REGION Network 164
   RUNG wire#powerrail
      Contact( "Carrier_27_Status.8" )
      Coil( "EMS".Carrier[27].SDC_IN.CrashDetectStatus )
   END_RUNG
   // the same network as SCL:
   "EMS".Carrier[27].SDC_IN.CrashDetectStatus := "Carrier_27_Status.8";
END_REGION

REGION Network 165
   RUNG wire#powerrail
      Contact( "Carrier_27_Status.9" )
      Coil( "EMS".Carrier[27].SDC_IN.EncoderCommFault )
   END_RUNG
   // the same network as SCL:
   "EMS".Carrier[27].SDC_IN.EncoderCommFault := "Carrier_27_Status.9";
END_REGION

REGION Network 166
   RUNG wire#powerrail
      Contact( "Carrier_27_Status.10" )
      Coil( "EMS".Carrier[27].SDC_IN.DriveCommFault )
   END_RUNG
   // the same network as SCL:
   "EMS".Carrier[27].SDC_IN.DriveCommFault := "Carrier_27_Status.10";
END_REGION

REGION Network 167
   RUNG wire#powerrail
      Contact( "Carrier_27_Status.11" )
      Coil( "EMS".Carrier[27].SDC_IN.HMICommFault )
   END_RUNG
   // the same network as SCL:
   "EMS".Carrier[27].SDC_IN.HMICommFault := "Carrier_27_Status.11";
END_REGION

REGION Network 168
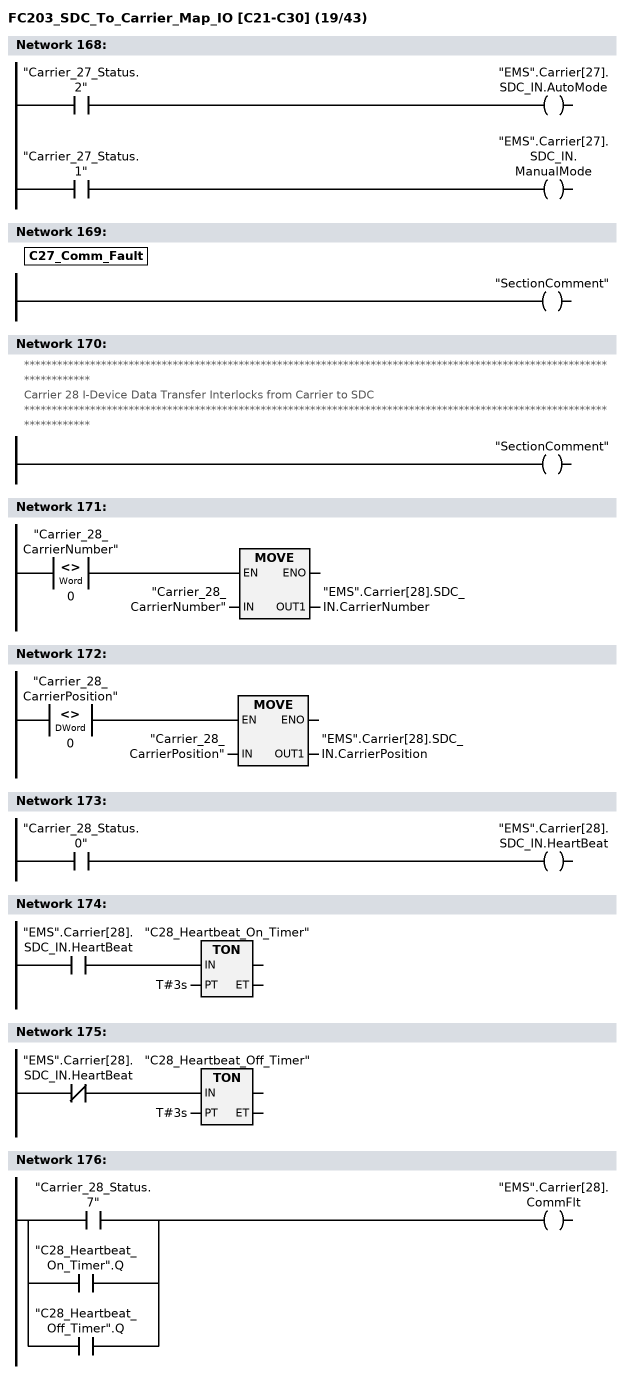
   RUNG wire#powerrail
      Contact( "Carrier_27_Status.2" )
      Coil( "EMS".Carrier[27].SDC_IN.AutoMode )
   END_RUNG
   RUNG wire#powerrail
      Contact( "Carrier_27_Status.1" )
      Coil( "EMS".Carrier[27].SDC_IN.ManualMode )
   END_RUNG
   // the same network as SCL:
   "EMS".Carrier[27].SDC_IN.AutoMode := "Carrier_27_Status.2";
   "EMS".Carrier[27].SDC_IN.ManualMode := "Carrier_27_Status.1";
END_REGION

REGION Network 169
   Label( C27_Comm_Fault )
   RUNG wire#powerrail
      Coil( "SectionComment" )
   END_RUNG
   // the same network as SCL:
   C27_Comm_Fault:
   "SectionComment" := TRUE;
END_REGION

REGION Network 170
   // **********************************************************************************************************************
   // 
   // Carrier 28 I-Device Data Transfer Interlocks from Carrier to SDC
   // 
   // **********************************************************************************************************************
   RUNG wire#powerrail
      Coil( "SectionComment" )
   END_RUNG
   // the same network as SCL:
   "SectionComment" := TRUE;
END_REGION

REGION Network 171
   RUNG wire#powerrail
      { S7_Templates := "SrcType := Word" } NE_Contact(in1 := "Carrier_28_CarrierNumber", in2 := 0)
      Move(in := "Carrier_28_CarrierNumber", out1 => "EMS".Carrier[28].SDC_IN.CarrierNumber)
   END_RUNG
   // the same network as SCL:
   IF "Carrier_28_CarrierNumber" <> 0 THEN
       "EMS".Carrier[28].SDC_IN.CarrierNumber := "Carrier_28_CarrierNumber";
   END_IF;
END_REGION

REGION Network 172
   RUNG wire#powerrail
      { S7_Templates := "SrcType := DWord" } NE_Contact(in1 := "Carrier_28_CarrierPosition", in2 := 0)
      Move(in := "Carrier_28_CarrierPosition", out1 => "EMS".Carrier[28].SDC_IN.CarrierPosition)
   END_RUNG
   // the same network as SCL:
   IF "Carrier_28_CarrierPosition" <> 0 THEN
       "EMS".Carrier[28].SDC_IN.CarrierPosition := "Carrier_28_CarrierPosition";
   END_IF;
END_REGION

REGION Network 173
   RUNG wire#powerrail
      Contact( "Carrier_28_Status.0" )
      Coil( "EMS".Carrier[28].SDC_IN.HeartBeat )
   END_RUNG
   // the same network as SCL:
   "EMS".Carrier[28].SDC_IN.HeartBeat := "Carrier_28_Status.0";
END_REGION

REGION Network 174
   "C28_Heartbeat_On_Timer".TON(IN := "EMS".Carrier[28].SDC_IN.HeartBeat, PT := T#3s);
END_REGION

REGION Network 175
   "C28_Heartbeat_Off_Timer".TON(IN := NOT "EMS".Carrier[28].SDC_IN.HeartBeat, PT := T#3s);
END_REGION

REGION Network 176
   RUNG wire#powerrail
      Contact( "Carrier_28_Status.7" )
      wire#w1
      Coil( "EMS".Carrier[28].CommFlt )
   END_RUNG
   RUNG wire#powerrail
      Contact( "C28_Heartbeat_On_Timer".Q )
   END_RUNG wire#w1
   RUNG wire#powerrail
      Contact( "C28_Heartbeat_Off_Timer".Q )
   END_RUNG wire#w1
   // the same network as SCL:
   "EMS".Carrier[28].CommFlt := "Carrier_28_Status.7" OR "C28_Heartbeat_On_Timer".Q OR "C28_Heartbeat_Off_Timer".Q;
END_REGION

REGION Network 177
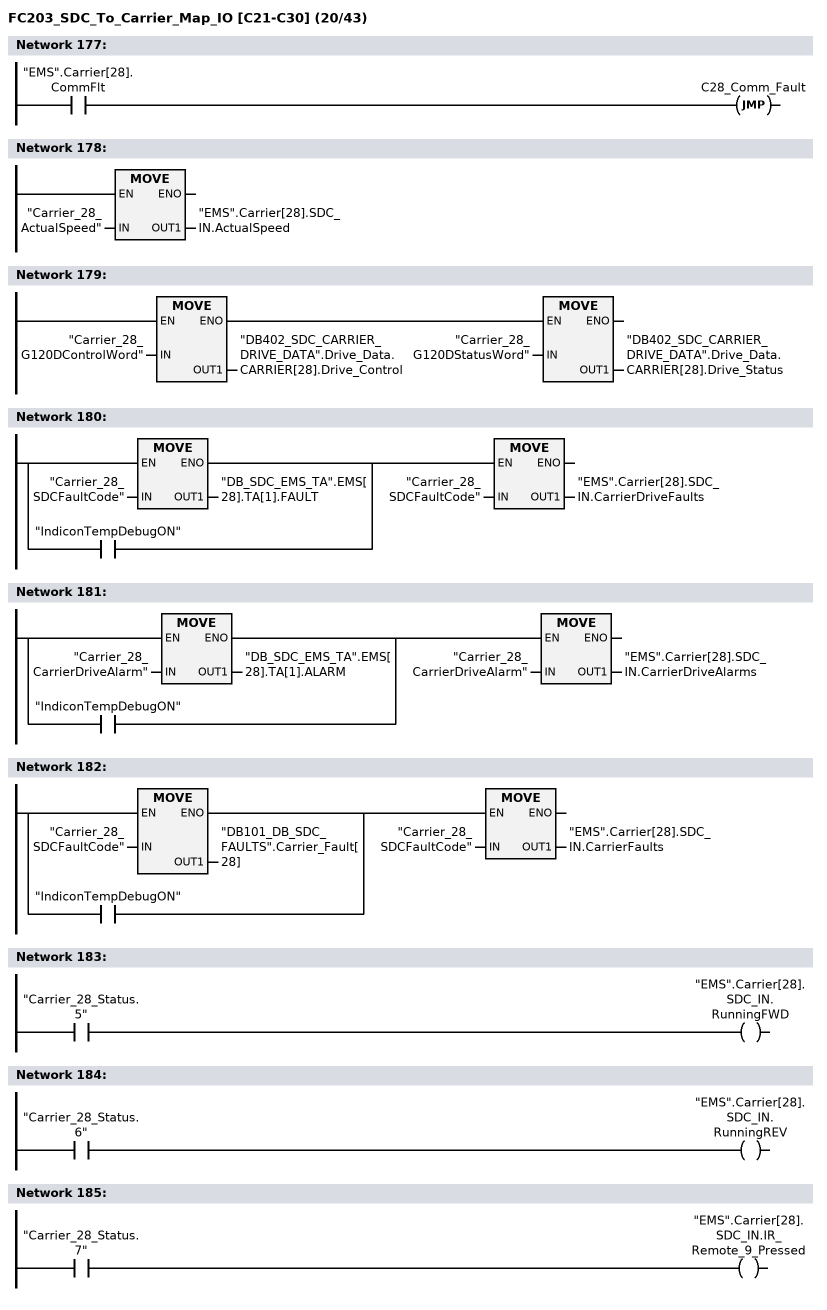
   RUNG wire#powerrail
      Contact( "EMS".Carrier[28].CommFlt )
      JumpCoil( C28_Comm_Fault )
   END_RUNG
   // the same network as SCL:
   IF "EMS".Carrier[28].CommFlt THEN GOTO C28_Comm_Fault; END_IF;
END_REGION

REGION Network 178
   RUNG wire#powerrail
      Move(in := "Carrier_28_ActualSpeed", out1 => "EMS".Carrier[28].SDC_IN.ActualSpeed)
   END_RUNG
   // the same network as SCL:
   "EMS".Carrier[28].SDC_IN.ActualSpeed := "Carrier_28_ActualSpeed";
END_REGION

REGION Network 179
   RUNG wire#powerrail
      Move(in := "Carrier_28_G120DControlWord", out1 => "DB402_SDC_CARRIER_DRIVE_DATA".Drive_Data.CARRIER[28].Drive_Control)
      Move(in := "Carrier_28_G120DStatusWord", out1 => "DB402_SDC_CARRIER_DRIVE_DATA".Drive_Data.CARRIER[28].Drive_Status)
   END_RUNG
   // the same network as SCL:
   "DB402_SDC_CARRIER_DRIVE_DATA".Drive_Data.CARRIER[28].Drive_Control := "Carrier_28_G120DControlWord";
   "DB402_SDC_CARRIER_DRIVE_DATA".Drive_Data.CARRIER[28].Drive_Status := "Carrier_28_G120DStatusWord";
END_REGION

REGION Network 180
   RUNG wire#powerrail
      Move(in := "Carrier_28_SDCFaultCode", out1 => "DB_SDC_EMS_TA".EMS[28].TA[1].FAULT)
      wire#w1
      Move(in := "Carrier_28_SDCFaultCode", out1 => "EMS".Carrier[28].SDC_IN.CarrierDriveFaults)
   END_RUNG
   RUNG wire#powerrail
      Contact( "IndiconTempDebugON" )
   END_RUNG wire#w1
   // the same network as SCL:
   "DB_SDC_EMS_TA".EMS[28].TA[1].FAULT := "Carrier_28_SDCFaultCode";
   IF TRUE OR "IndiconTempDebugON" THEN
       "EMS".Carrier[28].SDC_IN.CarrierDriveFaults := "Carrier_28_SDCFaultCode";
   END_IF;
END_REGION

REGION Network 181
   RUNG wire#powerrail
      Move(in := "Carrier_28_CarrierDriveAlarm", out1 => "DB_SDC_EMS_TA".EMS[28].TA[1].ALARM)
      wire#w1
      Move(in := "Carrier_28_CarrierDriveAlarm", out1 => "EMS".Carrier[28].SDC_IN.CarrierDriveAlarms)
   END_RUNG
   RUNG wire#powerrail
      Contact( "IndiconTempDebugON" )
   END_RUNG wire#w1
   // the same network as SCL:
   "DB_SDC_EMS_TA".EMS[28].TA[1].ALARM := "Carrier_28_CarrierDriveAlarm";
   IF TRUE OR "IndiconTempDebugON" THEN
       "EMS".Carrier[28].SDC_IN.CarrierDriveAlarms := "Carrier_28_CarrierDriveAlarm";
   END_IF;
END_REGION

REGION Network 182
   RUNG wire#powerrail
      Move(in := "Carrier_28_SDCFaultCode", out1 => "DB101_DB_SDC_FAULTS".Carrier_Fault[28])
      wire#w1
      Move(in := "Carrier_28_SDCFaultCode", out1 => "EMS".Carrier[28].SDC_IN.CarrierFaults)
   END_RUNG
   RUNG wire#powerrail
      Contact( "IndiconTempDebugON" )
   END_RUNG wire#w1
   // the same network as SCL:
   "DB101_DB_SDC_FAULTS".Carrier_Fault[28] := "Carrier_28_SDCFaultCode";
   IF TRUE OR "IndiconTempDebugON" THEN
       "EMS".Carrier[28].SDC_IN.CarrierFaults := "Carrier_28_SDCFaultCode";
   END_IF;
END_REGION

REGION Network 183
   RUNG wire#powerrail
      Contact( "Carrier_28_Status.5" )
      Coil( "EMS".Carrier[28].SDC_IN.RunningFWD )
   END_RUNG
   // the same network as SCL:
   "EMS".Carrier[28].SDC_IN.RunningFWD := "Carrier_28_Status.5";
END_REGION

REGION Network 184
   RUNG wire#powerrail
      Contact( "Carrier_28_Status.6" )
      Coil( "EMS".Carrier[28].SDC_IN.RunningREV )
   END_RUNG
   // the same network as SCL:
   "EMS".Carrier[28].SDC_IN.RunningREV := "Carrier_28_Status.6";
END_REGION

REGION Network 185
   RUNG wire#powerrail
      Contact( "Carrier_28_Status.7" )
      Coil( "EMS".Carrier[28].SDC_IN.IR_Remote_9_Pressed )
   END_RUNG
   // the same network as SCL:
   "EMS".Carrier[28].SDC_IN.IR_Remote_9_Pressed := "Carrier_28_Status.7";
END_REGION

REGION Network 186
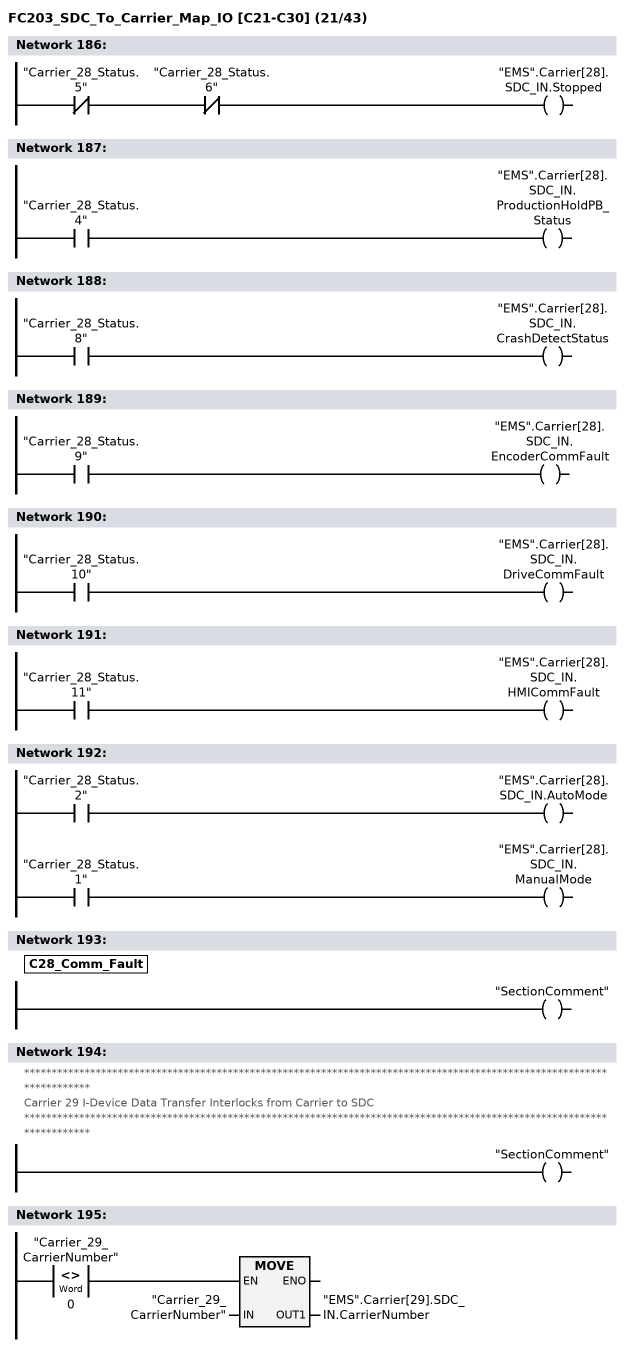
   RUNG wire#powerrail
      I_Contact( "Carrier_28_Status.5" )
      I_Contact( "Carrier_28_Status.6" )
      Coil( "EMS".Carrier[28].SDC_IN.Stopped )
   END_RUNG
   // the same network as SCL:
   "EMS".Carrier[28].SDC_IN.Stopped := NOT "Carrier_28_Status.5" AND NOT "Carrier_28_Status.6";
END_REGION

REGION Network 187
   RUNG wire#powerrail
      Contact( "Carrier_28_Status.4" )
      Coil( "EMS".Carrier[28].SDC_IN.ProductionHoldPB_Status )
   END_RUNG
   // the same network as SCL:
   "EMS".Carrier[28].SDC_IN.ProductionHoldPB_Status := "Carrier_28_Status.4";
END_REGION

REGION Network 188
   RUNG wire#powerrail
      Contact( "Carrier_28_Status.8" )
      Coil( "EMS".Carrier[28].SDC_IN.CrashDetectStatus )
   END_RUNG
   // the same network as SCL:
   "EMS".Carrier[28].SDC_IN.CrashDetectStatus := "Carrier_28_Status.8";
END_REGION

REGION Network 189
   RUNG wire#powerrail
      Contact( "Carrier_28_Status.9" )
      Coil( "EMS".Carrier[28].SDC_IN.EncoderCommFault )
   END_RUNG
   // the same network as SCL:
   "EMS".Carrier[28].SDC_IN.EncoderCommFault := "Carrier_28_Status.9";
END_REGION

REGION Network 190
   RUNG wire#powerrail
      Contact( "Carrier_28_Status.10" )
      Coil( "EMS".Carrier[28].SDC_IN.DriveCommFault )
   END_RUNG
   // the same network as SCL:
   "EMS".Carrier[28].SDC_IN.DriveCommFault := "Carrier_28_Status.10";
END_REGION

REGION Network 191
   RUNG wire#powerrail
      Contact( "Carrier_28_Status.11" )
      Coil( "EMS".Carrier[28].SDC_IN.HMICommFault )
   END_RUNG
   // the same network as SCL:
   "EMS".Carrier[28].SDC_IN.HMICommFault := "Carrier_28_Status.11";
END_REGION

REGION Network 192
   RUNG wire#powerrail
      Contact( "Carrier_28_Status.2" )
      Coil( "EMS".Carrier[28].SDC_IN.AutoMode )
   END_RUNG
   RUNG wire#powerrail
      Contact( "Carrier_28_Status.1" )
      Coil( "EMS".Carrier[28].SDC_IN.ManualMode )
   END_RUNG
   // the same network as SCL:
   "EMS".Carrier[28].SDC_IN.AutoMode := "Carrier_28_Status.2";
   "EMS".Carrier[28].SDC_IN.ManualMode := "Carrier_28_Status.1";
END_REGION

REGION Network 193
   Label( C28_Comm_Fault )
   RUNG wire#powerrail
      Coil( "SectionComment" )
   END_RUNG
   // the same network as SCL:
   C28_Comm_Fault:
   "SectionComment" := TRUE;
END_REGION

REGION Network 194
   // **********************************************************************************************************************
   // 
   // Carrier 29 I-Device Data Transfer Interlocks from Carrier to SDC
   // 
   // **********************************************************************************************************************
   RUNG wire#powerrail
      Coil( "SectionComment" )
   END_RUNG
   // the same network as SCL:
   "SectionComment" := TRUE;
END_REGION

REGION Network 195
   RUNG wire#powerrail
      { S7_Templates := "SrcType := Word" } NE_Contact(in1 := "Carrier_29_CarrierNumber", in2 := 0)
      Move(in := "Carrier_29_CarrierNumber", out1 => "EMS".Carrier[29].SDC_IN.CarrierNumber)
   END_RUNG
   // the same network as SCL:
   IF "Carrier_29_CarrierNumber" <> 0 THEN
       "EMS".Carrier[29].SDC_IN.CarrierNumber := "Carrier_29_CarrierNumber";
   END_IF;
END_REGION

REGION Network 196
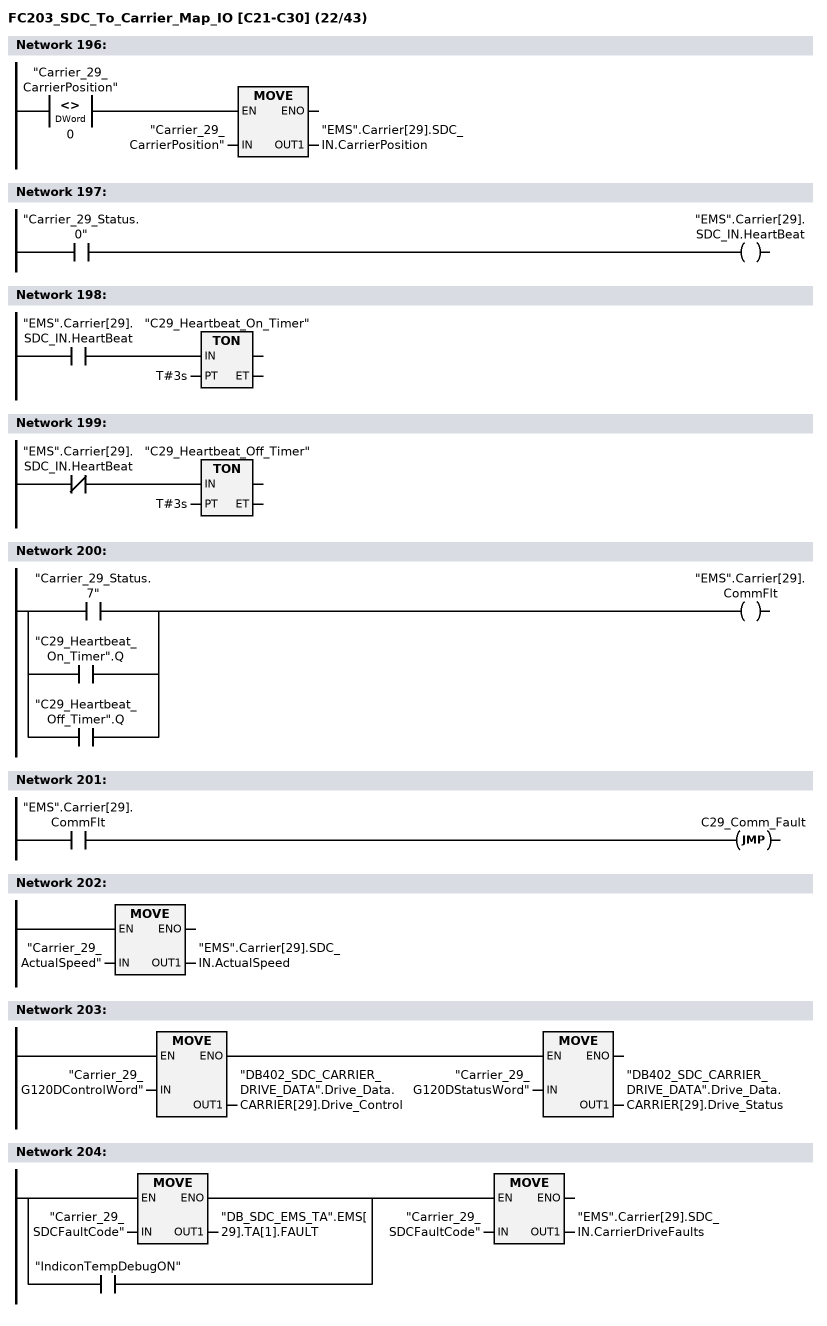
   RUNG wire#powerrail
      { S7_Templates := "SrcType := DWord" } NE_Contact(in1 := "Carrier_29_CarrierPosition", in2 := 0)
      Move(in := "Carrier_29_CarrierPosition", out1 => "EMS".Carrier[29].SDC_IN.CarrierPosition)
   END_RUNG
   // the same network as SCL:
   IF "Carrier_29_CarrierPosition" <> 0 THEN
       "EMS".Carrier[29].SDC_IN.CarrierPosition := "Carrier_29_CarrierPosition";
   END_IF;
END_REGION

REGION Network 197
   RUNG wire#powerrail
      Contact( "Carrier_29_Status.0" )
      Coil( "EMS".Carrier[29].SDC_IN.HeartBeat )
   END_RUNG
   // the same network as SCL:
   "EMS".Carrier[29].SDC_IN.HeartBeat := "Carrier_29_Status.0";
END_REGION

REGION Network 198
   "C29_Heartbeat_On_Timer".TON(IN := "EMS".Carrier[29].SDC_IN.HeartBeat, PT := T#3s);
END_REGION

REGION Network 199
   "C29_Heartbeat_Off_Timer".TON(IN := NOT "EMS".Carrier[29].SDC_IN.HeartBeat, PT := T#3s);
END_REGION

REGION Network 200
   RUNG wire#powerrail
      Contact( "Carrier_29_Status.7" )
      wire#w1
      Coil( "EMS".Carrier[29].CommFlt )
   END_RUNG
   RUNG wire#powerrail
      Contact( "C29_Heartbeat_On_Timer".Q )
   END_RUNG wire#w1
   RUNG wire#powerrail
      Contact( "C29_Heartbeat_Off_Timer".Q )
   END_RUNG wire#w1
   // the same network as SCL:
   "EMS".Carrier[29].CommFlt := "Carrier_29_Status.7" OR "C29_Heartbeat_On_Timer".Q OR "C29_Heartbeat_Off_Timer".Q;
END_REGION

REGION Network 201
   RUNG wire#powerrail
      Contact( "EMS".Carrier[29].CommFlt )
      JumpCoil( C29_Comm_Fault )
   END_RUNG
   // the same network as SCL:
   IF "EMS".Carrier[29].CommFlt THEN GOTO C29_Comm_Fault; END_IF;
END_REGION

REGION Network 202
   RUNG wire#powerrail
      Move(in := "Carrier_29_ActualSpeed", out1 => "EMS".Carrier[29].SDC_IN.ActualSpeed)
   END_RUNG
   // the same network as SCL:
   "EMS".Carrier[29].SDC_IN.ActualSpeed := "Carrier_29_ActualSpeed";
END_REGION

REGION Network 203
   RUNG wire#powerrail
      Move(in := "Carrier_29_G120DControlWord", out1 => "DB402_SDC_CARRIER_DRIVE_DATA".Drive_Data.CARRIER[29].Drive_Control)
      Move(in := "Carrier_29_G120DStatusWord", out1 => "DB402_SDC_CARRIER_DRIVE_DATA".Drive_Data.CARRIER[29].Drive_Status)
   END_RUNG
   // the same network as SCL:
   "DB402_SDC_CARRIER_DRIVE_DATA".Drive_Data.CARRIER[29].Drive_Control := "Carrier_29_G120DControlWord";
   "DB402_SDC_CARRIER_DRIVE_DATA".Drive_Data.CARRIER[29].Drive_Status := "Carrier_29_G120DStatusWord";
END_REGION

REGION Network 204
   RUNG wire#powerrail
      Move(in := "Carrier_29_SDCFaultCode", out1 => "DB_SDC_EMS_TA".EMS[29].TA[1].FAULT)
      wire#w1
      Move(in := "Carrier_29_SDCFaultCode", out1 => "EMS".Carrier[29].SDC_IN.CarrierDriveFaults)
   END_RUNG
   RUNG wire#powerrail
      Contact( "IndiconTempDebugON" )
   END_RUNG wire#w1
   // the same network as SCL:
   "DB_SDC_EMS_TA".EMS[29].TA[1].FAULT := "Carrier_29_SDCFaultCode";
   IF TRUE OR "IndiconTempDebugON" THEN
       "EMS".Carrier[29].SDC_IN.CarrierDriveFaults := "Carrier_29_SDCFaultCode";
   END_IF;
END_REGION

REGION Network 205
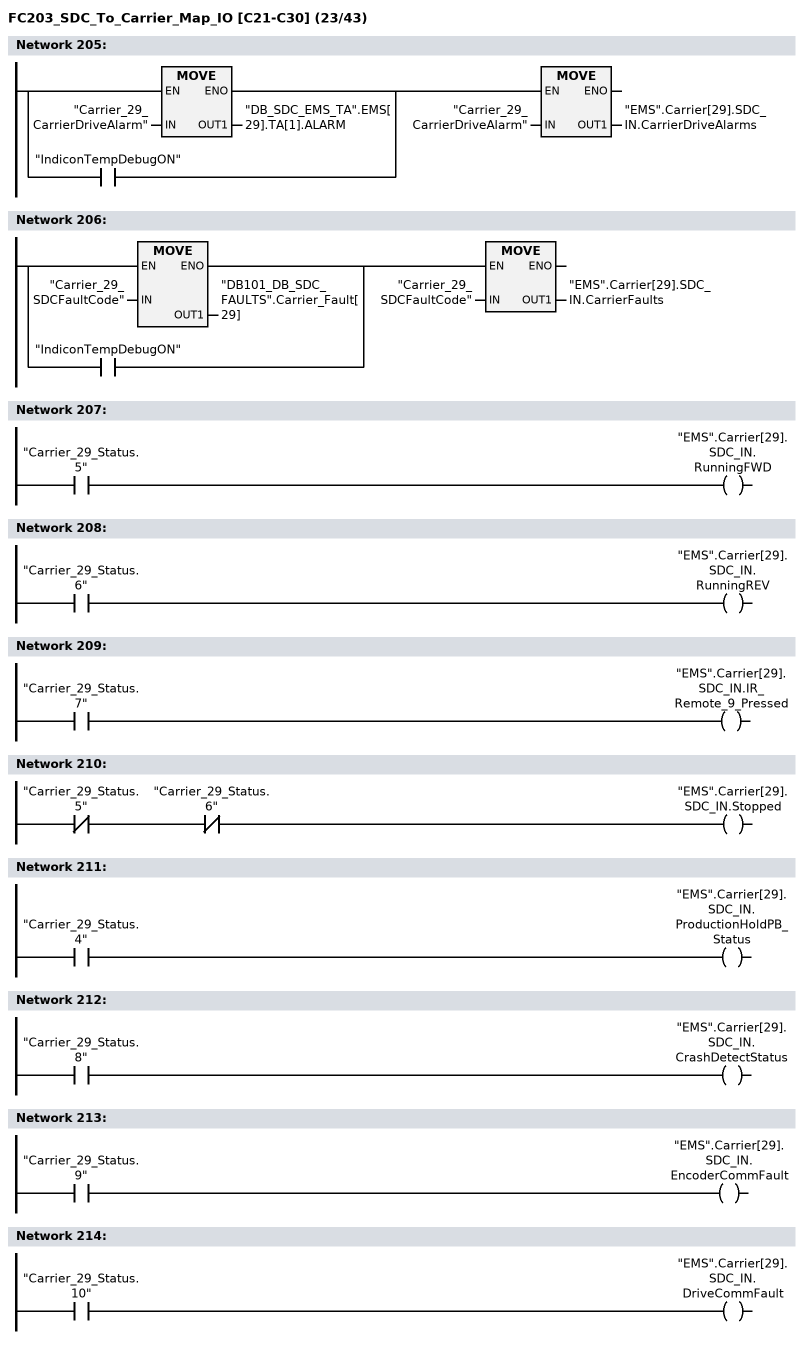
   RUNG wire#powerrail
      Move(in := "Carrier_29_CarrierDriveAlarm", out1 => "DB_SDC_EMS_TA".EMS[29].TA[1].ALARM)
      wire#w1
      Move(in := "Carrier_29_CarrierDriveAlarm", out1 => "EMS".Carrier[29].SDC_IN.CarrierDriveAlarms)
   END_RUNG
   RUNG wire#powerrail
      Contact( "IndiconTempDebugON" )
   END_RUNG wire#w1
   // the same network as SCL:
   "DB_SDC_EMS_TA".EMS[29].TA[1].ALARM := "Carrier_29_CarrierDriveAlarm";
   IF TRUE OR "IndiconTempDebugON" THEN
       "EMS".Carrier[29].SDC_IN.CarrierDriveAlarms := "Carrier_29_CarrierDriveAlarm";
   END_IF;
END_REGION

REGION Network 206
   RUNG wire#powerrail
      Move(in := "Carrier_29_SDCFaultCode", out1 => "DB101_DB_SDC_FAULTS".Carrier_Fault[29])
      wire#w1
      Move(in := "Carrier_29_SDCFaultCode", out1 => "EMS".Carrier[29].SDC_IN.CarrierFaults)
   END_RUNG
   RUNG wire#powerrail
      Contact( "IndiconTempDebugON" )
   END_RUNG wire#w1
   // the same network as SCL:
   "DB101_DB_SDC_FAULTS".Carrier_Fault[29] := "Carrier_29_SDCFaultCode";
   IF TRUE OR "IndiconTempDebugON" THEN
       "EMS".Carrier[29].SDC_IN.CarrierFaults := "Carrier_29_SDCFaultCode";
   END_IF;
END_REGION

REGION Network 207
   RUNG wire#powerrail
      Contact( "Carrier_29_Status.5" )
      Coil( "EMS".Carrier[29].SDC_IN.RunningFWD )
   END_RUNG
   // the same network as SCL:
   "EMS".Carrier[29].SDC_IN.RunningFWD := "Carrier_29_Status.5";
END_REGION

REGION Network 208
   RUNG wire#powerrail
      Contact( "Carrier_29_Status.6" )
      Coil( "EMS".Carrier[29].SDC_IN.RunningREV )
   END_RUNG
   // the same network as SCL:
   "EMS".Carrier[29].SDC_IN.RunningREV := "Carrier_29_Status.6";
END_REGION

REGION Network 209
   RUNG wire#powerrail
      Contact( "Carrier_29_Status.7" )
      Coil( "EMS".Carrier[29].SDC_IN.IR_Remote_9_Pressed )
   END_RUNG
   // the same network as SCL:
   "EMS".Carrier[29].SDC_IN.IR_Remote_9_Pressed := "Carrier_29_Status.7";
END_REGION

REGION Network 210
   RUNG wire#powerrail
      I_Contact( "Carrier_29_Status.5" )
      I_Contact( "Carrier_29_Status.6" )
      Coil( "EMS".Carrier[29].SDC_IN.Stopped )
   END_RUNG
   // the same network as SCL:
   "EMS".Carrier[29].SDC_IN.Stopped := NOT "Carrier_29_Status.5" AND NOT "Carrier_29_Status.6";
END_REGION

REGION Network 211
   RUNG wire#powerrail
      Contact( "Carrier_29_Status.4" )
      Coil( "EMS".Carrier[29].SDC_IN.ProductionHoldPB_Status )
   END_RUNG
   // the same network as SCL:
   "EMS".Carrier[29].SDC_IN.ProductionHoldPB_Status := "Carrier_29_Status.4";
END_REGION

REGION Network 212
   RUNG wire#powerrail
      Contact( "Carrier_29_Status.8" )
      Coil( "EMS".Carrier[29].SDC_IN.CrashDetectStatus )
   END_RUNG
   // the same network as SCL:
   "EMS".Carrier[29].SDC_IN.CrashDetectStatus := "Carrier_29_Status.8";
END_REGION

REGION Network 213
   RUNG wire#powerrail
      Contact( "Carrier_29_Status.9" )
      Coil( "EMS".Carrier[29].SDC_IN.EncoderCommFault )
   END_RUNG
   // the same network as SCL:
   "EMS".Carrier[29].SDC_IN.EncoderCommFault := "Carrier_29_Status.9";
END_REGION

REGION Network 214
   RUNG wire#powerrail
      Contact( "Carrier_29_Status.10" )
      Coil( "EMS".Carrier[29].SDC_IN.DriveCommFault )
   END_RUNG
   // the same network as SCL:
   "EMS".Carrier[29].SDC_IN.DriveCommFault := "Carrier_29_Status.10";
END_REGION

REGION Network 215
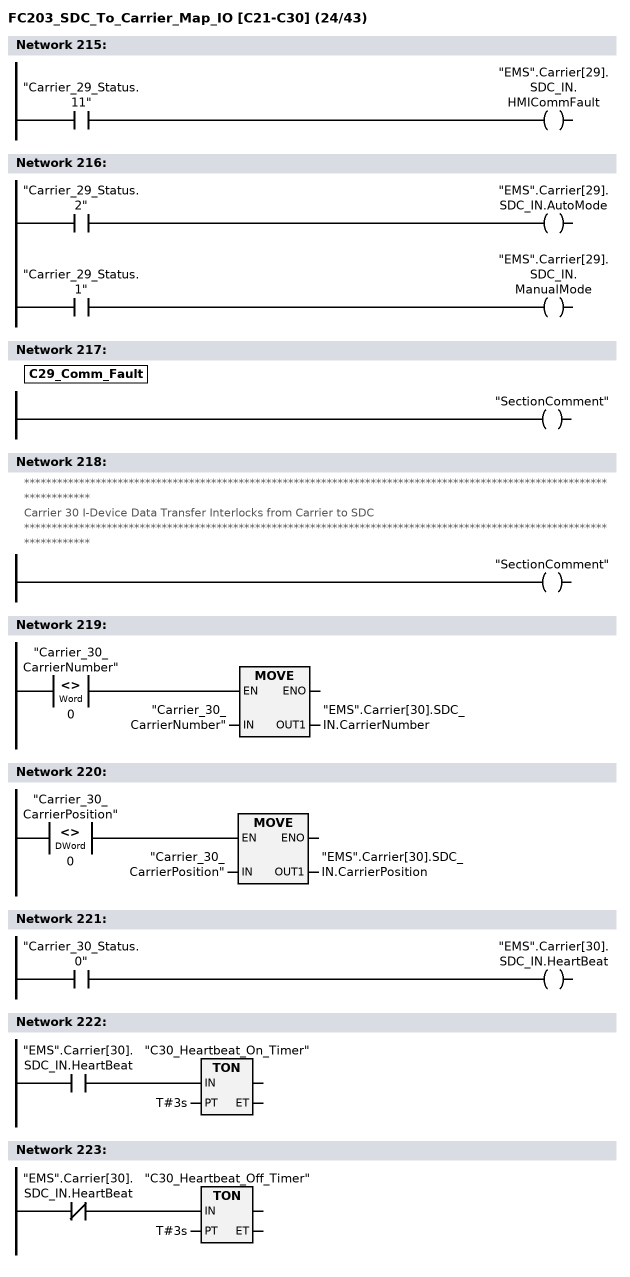
   RUNG wire#powerrail
      Contact( "Carrier_29_Status.11" )
      Coil( "EMS".Carrier[29].SDC_IN.HMICommFault )
   END_RUNG
   // the same network as SCL:
   "EMS".Carrier[29].SDC_IN.HMICommFault := "Carrier_29_Status.11";
END_REGION

REGION Network 216
   RUNG wire#powerrail
      Contact( "Carrier_29_Status.2" )
      Coil( "EMS".Carrier[29].SDC_IN.AutoMode )
   END_RUNG
   RUNG wire#powerrail
      Contact( "Carrier_29_Status.1" )
      Coil( "EMS".Carrier[29].SDC_IN.ManualMode )
   END_RUNG
   // the same network as SCL:
   "EMS".Carrier[29].SDC_IN.AutoMode := "Carrier_29_Status.2";
   "EMS".Carrier[29].SDC_IN.ManualMode := "Carrier_29_Status.1";
END_REGION

REGION Network 217
   Label( C29_Comm_Fault )
   RUNG wire#powerrail
      Coil( "SectionComment" )
   END_RUNG
   // the same network as SCL:
   C29_Comm_Fault:
   "SectionComment" := TRUE;
END_REGION

REGION Network 218
   // **********************************************************************************************************************
   // 
   // Carrier 30 I-Device Data Transfer Interlocks from Carrier to SDC
   // 
   // **********************************************************************************************************************
   RUNG wire#powerrail
      Coil( "SectionComment" )
   END_RUNG
   // the same network as SCL:
   "SectionComment" := TRUE;
END_REGION

REGION Network 219
   RUNG wire#powerrail
      { S7_Templates := "SrcType := Word" } NE_Contact(in1 := "Carrier_30_CarrierNumber", in2 := 0)
      Move(in := "Carrier_30_CarrierNumber", out1 => "EMS".Carrier[30].SDC_IN.CarrierNumber)
   END_RUNG
   // the same network as SCL:
   IF "Carrier_30_CarrierNumber" <> 0 THEN
       "EMS".Carrier[30].SDC_IN.CarrierNumber := "Carrier_30_CarrierNumber";
   END_IF;
END_REGION

REGION Network 220
   RUNG wire#powerrail
      { S7_Templates := "SrcType := DWord" } NE_Contact(in1 := "Carrier_30_CarrierPosition", in2 := 0)
      Move(in := "Carrier_30_CarrierPosition", out1 => "EMS".Carrier[30].SDC_IN.CarrierPosition)
   END_RUNG
   // the same network as SCL:
   IF "Carrier_30_CarrierPosition" <> 0 THEN
       "EMS".Carrier[30].SDC_IN.CarrierPosition := "Carrier_30_CarrierPosition";
   END_IF;
END_REGION

REGION Network 221
   RUNG wire#powerrail
      Contact( "Carrier_30_Status.0" )
      Coil( "EMS".Carrier[30].SDC_IN.HeartBeat )
   END_RUNG
   // the same network as SCL:
   "EMS".Carrier[30].SDC_IN.HeartBeat := "Carrier_30_Status.0";
END_REGION

REGION Network 222
   "C30_Heartbeat_On_Timer".TON(IN := "EMS".Carrier[30].SDC_IN.HeartBeat, PT := T#3s);
END_REGION

REGION Network 223
   "C30_Heartbeat_Off_Timer".TON(IN := NOT "EMS".Carrier[30].SDC_IN.HeartBeat, PT := T#3s);
END_REGION

REGION Network 224
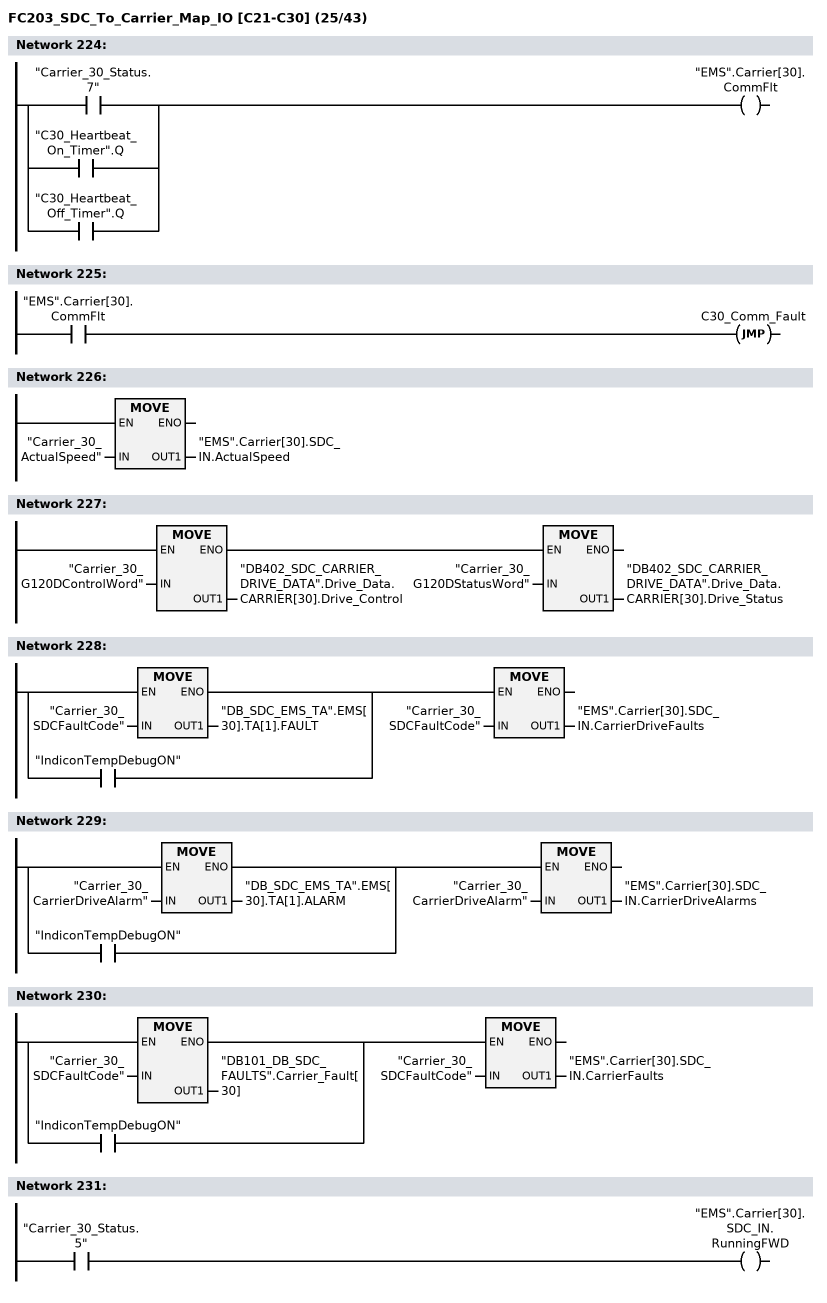
   RUNG wire#powerrail
      Contact( "Carrier_30_Status.7" )
      wire#w1
      Coil( "EMS".Carrier[30].CommFlt )
   END_RUNG
   RUNG wire#powerrail
      Contact( "C30_Heartbeat_On_Timer".Q )
   END_RUNG wire#w1
   RUNG wire#powerrail
      Contact( "C30_Heartbeat_Off_Timer".Q )
   END_RUNG wire#w1
   // the same network as SCL:
   "EMS".Carrier[30].CommFlt := "Carrier_30_Status.7" OR "C30_Heartbeat_On_Timer".Q OR "C30_Heartbeat_Off_Timer".Q;
END_REGION

REGION Network 225
   RUNG wire#powerrail
      Contact( "EMS".Carrier[30].CommFlt )
      JumpCoil( C30_Comm_Fault )
   END_RUNG
   // the same network as SCL:
   IF "EMS".Carrier[30].CommFlt THEN GOTO C30_Comm_Fault; END_IF;
END_REGION

REGION Network 226
   RUNG wire#powerrail
      Move(in := "Carrier_30_ActualSpeed", out1 => "EMS".Carrier[30].SDC_IN.ActualSpeed)
   END_RUNG
   // the same network as SCL:
   "EMS".Carrier[30].SDC_IN.ActualSpeed := "Carrier_30_ActualSpeed";
END_REGION

REGION Network 227
   RUNG wire#powerrail
      Move(in := "Carrier_30_G120DControlWord", out1 => "DB402_SDC_CARRIER_DRIVE_DATA".Drive_Data.CARRIER[30].Drive_Control)
      Move(in := "Carrier_30_G120DStatusWord", out1 => "DB402_SDC_CARRIER_DRIVE_DATA".Drive_Data.CARRIER[30].Drive_Status)
   END_RUNG
   // the same network as SCL:
   "DB402_SDC_CARRIER_DRIVE_DATA".Drive_Data.CARRIER[30].Drive_Control := "Carrier_30_G120DControlWord";
   "DB402_SDC_CARRIER_DRIVE_DATA".Drive_Data.CARRIER[30].Drive_Status := "Carrier_30_G120DStatusWord";
END_REGION

REGION Network 228
   RUNG wire#powerrail
      Move(in := "Carrier_30_SDCFaultCode", out1 => "DB_SDC_EMS_TA".EMS[30].TA[1].FAULT)
      wire#w1
      Move(in := "Carrier_30_SDCFaultCode", out1 => "EMS".Carrier[30].SDC_IN.CarrierDriveFaults)
   END_RUNG
   RUNG wire#powerrail
      Contact( "IndiconTempDebugON" )
   END_RUNG wire#w1
   // the same network as SCL:
   "DB_SDC_EMS_TA".EMS[30].TA[1].FAULT := "Carrier_30_SDCFaultCode";
   IF TRUE OR "IndiconTempDebugON" THEN
       "EMS".Carrier[30].SDC_IN.CarrierDriveFaults := "Carrier_30_SDCFaultCode";
   END_IF;
END_REGION

REGION Network 229
   RUNG wire#powerrail
      Move(in := "Carrier_30_CarrierDriveAlarm", out1 => "DB_SDC_EMS_TA".EMS[30].TA[1].ALARM)
      wire#w1
      Move(in := "Carrier_30_CarrierDriveAlarm", out1 => "EMS".Carrier[30].SDC_IN.CarrierDriveAlarms)
   END_RUNG
   RUNG wire#powerrail
      Contact( "IndiconTempDebugON" )
   END_RUNG wire#w1
   // the same network as SCL:
   "DB_SDC_EMS_TA".EMS[30].TA[1].ALARM := "Carrier_30_CarrierDriveAlarm";
   IF TRUE OR "IndiconTempDebugON" THEN
       "EMS".Carrier[30].SDC_IN.CarrierDriveAlarms := "Carrier_30_CarrierDriveAlarm";
   END_IF;
END_REGION

REGION Network 230
   RUNG wire#powerrail
      Move(in := "Carrier_30_SDCFaultCode", out1 => "DB101_DB_SDC_FAULTS".Carrier_Fault[30])
      wire#w1
      Move(in := "Carrier_30_SDCFaultCode", out1 => "EMS".Carrier[30].SDC_IN.CarrierFaults)
   END_RUNG
   RUNG wire#powerrail
      Contact( "IndiconTempDebugON" )
   END_RUNG wire#w1
   // the same network as SCL:
   "DB101_DB_SDC_FAULTS".Carrier_Fault[30] := "Carrier_30_SDCFaultCode";
   IF TRUE OR "IndiconTempDebugON" THEN
       "EMS".Carrier[30].SDC_IN.CarrierFaults := "Carrier_30_SDCFaultCode";
   END_IF;
END_REGION

REGION Network 231
   RUNG wire#powerrail
      Contact( "Carrier_30_Status.5" )
      Coil( "EMS".Carrier[30].SDC_IN.RunningFWD )
   END_RUNG
   // the same network as SCL:
   "EMS".Carrier[30].SDC_IN.RunningFWD := "Carrier_30_Status.5";
END_REGION

REGION Network 232